screen "0012_Pump Setting" 1280x800, template "Navigation"
   on GenerateScreen: SetBit("DB613_Komponent_State_Read"); SetBit("DB608_PV_Metering_Read")
   Button "Button_1" at 133,154 size 561x639; TextOff 'Text'
   TextField "Text field_1" at 170,166 size 134x25; Text 'Pump enable:'
   TextField "Text field_2" at 170,199 size 128x25; Text 'Machine No.:'
   TextField "Text field_3" at 170,231 size 90x25; Text 'Daytank:'
   TextField "Text field_4" at 170,296 size 65x25; Text 'Name:'
   TextField "Text field_5" at 170,326 size 156x25; Text 'Pulse per. Liter:'
   TextField "Text field_7" at 170,357 size 196x25; Text 'Adjustm. time [ms]:'
   IOField "Pump_Pulse_Perliter" at 453,323 size 166x30; Authorization "User administration"; FormatPattern 99999.999
      ProcessValue <- "DB753_MeteringPump_Pump{0}_Pulse_per_liter"
   TextField "Text field_8" at 170,550 size 82x25; Text 'Control:'
   TextField "Text field_9" at 170,582 size 146x25; Text 'Feeding Pump:'
   TextField "Text field_10" at 170,617 size 114x25; Text 'Edge Filter:'
   TextField "Text field_11" at 170,652 size 181x25; Text 'Cooling / Heating:'
   TextField "Text field_12" at 170,687 size 192x25; Text 'Deselection Enable:'
   TextField "Text field_13" at 170,722 size 302x25; Text 'With min Temperature Release:'
   TextField "Text field_14" at 170,757 size 167x25; Text 'With flow factor:'
   IOField "I/O field_2" at 453,354 size 166x30; Authorization "User administration"; FormatPattern 99999.999
      ProcessValue <- "PN_FlowRate_Component{0}_FlowC_F_GeneralParameters_Data_Nachstellzeit"
   IOField "I/O field_3" at 453,385 size 166x30; Authorization "User administration"; FormatPattern 999.9
      ProcessValue <- "DB753_MeteringPump_Pump{0}_MaxFlowLiter"
   IOField "I/O field_4" at 551,196 size 69x30; Authorization "User administration"; FormatPattern 999
      ProcessValue <- "DB753_MeteringPump_Pump{0}_MachineNumber"
   IOField "I/O field_5" at 551,228 size 69x30; Authorization "User administration"; FormatPattern 9999
      ProcessValue <- "DB753_MeteringPump_Pump{0}_TankNo"
   Button "Check_Pump_Enable" at 575,161 size 45x30; TextOff 'Text'; PictureOff "download"; PictureList "Check_Uncheck"
      ProcessValue <- "DB753_MeteringPump_Pump{0}_Pump_Active"
      on Click: InvertBit("DB753_MeteringPump_Pump{0}_Pump_Active")
   Button "Check_Pump_WithFeedingPump" at 573,579 size 45x30; TextOff 'Text'; PictureOff "download"; PictureList "Check_Uncheck"
      ProcessValue <- "DB753_MeteringPump_Pump{0}_WithFeedPump"
      on Click: InvertBit("DB753_MeteringPump_Pump{0}_WithFeedPump")
   Button "Check_Pump_WithEdgeFilter" at 573,614 size 45x30; TextOff 'Text'; PictureOff "download"; PictureList "Check_Uncheck"
      ProcessValue <- "DB753_MeteringPump_Pump{0}_WithEdgeFilter"
      on Click: InvertBit("DB753_MeteringPump_Pump{0}_WithEdgeFilter")
   Button "Check_Pump_CoolingHeating" at 573,649 size 45x30; TextOff 'Text'; PictureOff "download"; PictureList "Check_Uncheck"
      ProcessValue <- "DB753_MeteringPump_Pump{0}_WithHeating"
      on Click: InvertBit("DB753_MeteringPump_Pump{0}_WithHeating")
   Button "Check_Pump_Deselection_Ena" at 573,684 size 45x30; TextOff 'Text'; PictureOff "download"; PictureList "Check_Uncheck"
      ProcessValue <- "DB753_MeteringPump_Pump{0}_PumDeselectionEnable"
      on Click: InvertBit("DB753_MeteringPump_Pump{0}_PumDeselectionEnable")
   Button "Check_Pump_WithMinTempRelease" at 573,719 size 45x30; TextOff 'Text'; PictureOff "download"; PictureList "Check_Uncheck"
      ProcessValue <- "DB753_MeteringPump_Pump{0}_WithMinTempRelease"
      on Click: InvertBit("DB753_MeteringPump_Pump{0}_WithMinTempRelease")
   Button "Check_Pump_WithFlowFactor" at 573,754 size 45x30; TextOff 'Text'; PictureOff "download"; PictureList "Check_Uncheck"
      ProcessValue <- "DB753_MeteringPump_Pump{0}_WithFlowFactor"
      on Click: InvertBit("DB753_MeteringPump_Pump{0}_WithFlowFactor")
   Button "b_Incress_Pump_Setting" at 785,104 size 46x32; TextOff 'Text'; PictureOff "right arrow"
      on Click: function_dd21b452("DB613_Komponent_State_ReadDeviceNo", 1); function_dd21b452("DB612_Tank_State.ReadDeviceNo", 1)
   Button "b_Decress_Pump_Setting" at 273,104 size 46x32; TextOff 'Text'; PictureOff "left arrow"
      on Click: function_b9b71300("DB613_Komponent_State_ReadDeviceNo", 1); function_b9b71300("DB612_Tank_State.ReadDeviceNo", 1)
   Button "b_Pump_Control" at 503,547 size 45x30; TextOff 'Text'; PictureOff "obeng"
      on Click: SetTag("Control", 1)
   Button "b_Pump_Feeding_Pump" at 503,579 size 45x30; TextOff 'Text'; PictureOff "obeng"
      on Click: SetTag("Control", 2)
      Visibility <- "DB753_MeteringPump_Pump{0}_WithFeedPump"
   Button "b_Pump_EdgeFilter" at 503,615 size 45x30; TextOff 'Text'; PictureOff "obeng"
      on Click: SetTag("Control", 3)
      Visibility <- "DB753_MeteringPump_Pump{0}_WithEdgeFilter"
   Button "b_Pump_CoolingHeating" at 503,651 size 45x30; TextOff 'Text'; PictureOff "obeng"
      on Click: SetTag("Control", 4)
      Visibility <- "DB753_MeteringPump_Pump{0}_WithHeating"
   IOField "I/O field_6" at 453,293 size 166x30; Authorization "User administration"; FormatPattern ??????????
      ProcessValue <- "DB753_MeteringPump_Pump{0}_Name"
   IOField "I/O field_7" at 382,261 size 236x30; Authorization "User administration"; FormatPattern ??????????
      ProcessValue <- "DB753_MeteringPump_Pump{0}_Name"
   IOField "I/O field_8" at 453,417 size 166x30; Authorization "User administration"; FormatPattern 999.9
      ProcessValue <- "DB753_MeteringPump_Pump{0}_MinFlowPercent"
   IOField "I/O field_9" at 453,449 size 166x30; Authorization "User administration"; FormatPattern 999.9
      ProcessValue <- "DB753_MeteringPump_Pump{0}_MaxFlowPercent"
   IOField "I/O field_10" at 453,479 size 166x30; Authorization "User administration"; FormatPattern 99999.99
      ProcessValue <- "DB613_Komponent_State_FlowPumpMin{0}"
   IOField "I/O field_11" at 453,511 size 166x30; Authorization "User administration"; FormatPattern 99999.99
      ProcessValue <- "DB613_Komponent_State_FlowPumpMax{0}"
   TextField "Text field_20" at 170,388 size 227x25; Text 'Pump quantity [l/min]:'
   TextField "Text field_21" at 170,420 size 142x25; Text 'Min. Flow[%]:'
   TextField "Text field_22" at 170,452 size 146x25; Text 'Max. Flow[%]:'
   TextField "Text field_23" at 170,482 size 154x25; Text 'Min. Flow[g/s]:'
   TextField "Text field_24" at 170,514 size 158x25; Text 'Max. Flow[g/s]:'
   IOField "I/O field_43" at 326,104 size 451x32; FormatPattern ????????????????????
      ProcessValue <- "DB753_MeteringPump_Pump{0}_Name"
      Appearance <- "DB702_Tank_Value_Tank{0}_Color"
   Button "Button_19" at 856,366 size 159x83; TextOff 'Text'; PictureOff "motor_2"; PictureList "pump"
      ProcessValue <- "DB613_Komponent_State_ReadDeviceNo"
      Visibility <- "DB753_MeteringPump_Pump{0}_Pump_Active"
   GraphicView "Graphic view_1" at 763,170 size 81x40; Picture "motor2"
      Visibility <- "DB753_MeteringPump_Pump{0}_WithFeedPump"
   GraphicView "Graphic view_2" at 715,254 size 125x120; Picture "heatHP"
      Visibility <- "DB753_MeteringPump_Pump{0}_WithHeating"
   GraphicView "Graphic view_5" at 1047,261 size 58x89; Picture "heatLP"
      Visibility <- "DB753_MeteringPump_Pump{0}_WithLPHeatExchanger"
   GraphicView "Graphic view_7" at 977,170 size 67x93; Picture "edgefilter"
      Visibility <- "DB753_MeteringPump_Pump{0}_WithEdgeFilter"
   GraphicView "Graphic view_9" at 1112,275 size 39x75; Picture "Graphic_14"
      Visibility <- "DB753_MeteringPump_Pump{0}_WithFischerValveLP"
   GraphicView "Graphic view_10" at 801,275 size 39x75; Picture "Graphic_14"
      Visibility <- "DB753_MeteringPump_Pump{0}_WithFischerValveHP"
   Button "Button_8" at 720,466 size 437x286; TextOff 'Text'
      Visibility <- "Control"
   TextField "Text field_15" at 742,497 size 169x30; Text 'Control Pump:'
      Visibility <- "Control"
   TextField "Text field_16" at 742,573 size 91x25; Text 'With FC :'
      Visibility <- "Control"
   TextField "Text field_17" at 742,617 size 104x25; Text 'Controlled'
      Visibility <- "Control"
   TextField "Text field_18" at 742,661 size 73x25; Text '2 Point'
      Visibility <- "Control"
   TextField "Text field_19" at 940,617 size 101x25; Text 'Regulated'
      Visibility <- "Control"
   Button "Check_Pump_ControlPump_WithFc" at 862,570 size 45x30; TextOff 'Text'; PictureOff "download"; PictureList "Check_Uncheck"
      ProcessValue <- "DB753_MeteringPump_Pump{0}_WithFC"
      Visibility <- "Control"
      on Click: InvertBit("DB753_MeteringPump_Pump{0}_WithFC")
   Button "Check_Pump_ControlPump_Controlled" at 862,614 size 45x30; TextOff 'Text'; PictureOff "download"; PictureList "Check_Uncheck"
      Visibility <- "Control"
      ProcessValue <- "DB753_MeteringPump_Pump{0}_WithFlowControl"
      on Click: InvertBit("DB753_MeteringPump_Pump{0}_WithFlowControl")
   Button "Check_Pump_ControlPump_2Point" at 862,658 size 45x30; TextOff 'Text'; PictureOff "download"; PictureList "Check_Uncheck"
      ProcessValue <- "DB753_MeteringPump_Pump{0}_With_2Point"
      Visibility <- "Control"
      on Click: InvertBit("DB753_MeteringPump_Pump{0}_With_2Point")
   Button "Check_Pump_ControlPump_Regulated" at 1057,614 size 45x30; TextOff 'Text'; PictureOff "download"; PictureList "Check_Uncheck"
      Visibility <- "Control"
      ProcessValue <- "DB753_MeteringPump_Pump{0}_WithoutFlowControl"
      on Click: InvertBit("DB753_MeteringPump_Pump{0}_WithoutFlowControl")
   Button "b_Pump_Close_ControlPump" at 1101,470 size 51x41; TextOff 'Text'; PictureOff "images (1)"
      Visibility <- "Control"
      on Click: SetTag("Control", 0)
   Button "Button_2" at 720,466 size 437x286; TextOff 'Text'
      Visibility <- "Control"
   TextField "Text field_6" at 758,496 size 173x30; Text 'Feeding Pump:'
      Visibility <- "Control"
   TextField "Text field_25" at 794,559 size 78x25; Text 'With FC'
      Visibility <- "Control"
   TextField "Text field_26" at 794,609 size 157x25; Text 'No pressure ctr.'
      Visibility <- "Control"
   TextField "Text field_27" at 794,657 size 72x25; Text 'Bypass'
      Visibility <- "Control"
   TextField "Text field_28" at 1023,559 size 125x25; Text 'Pressure ctr.'
      Visibility <- "Control"
   Button "Check_Pump_FP_WithFC" at 738,556 size 45x30; TextOff 'Text'; PictureOff "download"; PictureList "Check_Uncheck"
      Visibility <- "Control"
      on Click: InvertBit("DB751_auxiliaryDriveMetering_FeedingPump{0}_Config_WithFC")
      ProcessValue <- "DB751_auxiliaryDriveMetering_FeedingPump{0}_Config_WithFC"
   Button "Check_Pump_FP_NoPressCtr" at 738,606 size 45x30; TextOff 'Text'; PictureOff "download"; PictureList "Check_Uncheck"
      Visibility <- "Control"
      on Click: InvertBit("DB751_auxiliaryDriveMetering_FeedingPump{0}_Config_Without_PresControl")
      ProcessValue <- "DB751_auxiliaryDriveMetering_FeedingPump{0}_Config_Without_PresControl"
   Button "Check_Pump_FP_Bypass" at 738,654 size 45x30; TextOff 'Text'; PictureOff "download"; PictureList "Check_Uncheck"
      Visibility <- "Control"
      on Click: InvertBit("DB751_auxiliaryDriveMetering_FeedingPump{0}_Config_Bypass")
      ProcessValue <- "DB751_auxiliaryDriveMetering_FeedingPump{0}_Config_Bypass"
   Button "Check_Pump_FP_PressureCtr" at 963,556 size 45x30; TextOff 'Text'; PictureOff "download"; PictureList "Check_Uncheck"
      Visibility <- "Control"
      on Click: InvertBit("DB751_auxiliaryDriveMetering_FeedingPump{0}_Config_With_PresControl")
      ProcessValue <- "DB751_auxiliaryDriveMetering_FeedingPump{0}_Config_With_PresControl"
   Button "b_Close_Pump_FeddingPump" at 1101,469 size 51x41; TextOff 'Text'; PictureOff "images (1)"
      Visibility <- "Control"
      on Click: SetTag("Control", 0)
   TextField "Text field_29" at 794,705 size 154x25; Text 'Manual Switch?'
      Visibility <- "Control"
   Button "Check_Pump_FP_ManualSwtch?" at 738,702 size 45x30; TextOff 'Text'; PictureOff "download"; PictureList "Check_Uncheck"
      Visibility <- "Control"
      on Click: InvertBit("DB751_auxiliaryDriveMetering_FeedingPump{0}_Config_ManualSwitchON")
      ProcessValue <- "DB751_auxiliaryDriveMetering_FeedingPump{0}_Config_ManualSwitchON"
   TextField "Text field_30" at 1023,609 size 64x25; Text 'Filling'
      Visibility <- "Control"
   Button "Check-Pump_FP_Filling" at 963,606 size 45x30; TextOff 'Text'; PictureOff "download"; PictureList "Check_Uncheck"
      Visibility <- "Control"
      on Click: InvertBit("DB751_auxiliaryDriveMetering_FeedingPump{0}_Config_Filling")
      ProcessValue <- "DB751_auxiliaryDriveMetering_FeedingPump{0}_Config_Filling"
   Button "Button_11" at 720,466 size 437x286; TextOff 'Text'
      Visibility <- "Control"
   TextField "Text field_31" at 754,496 size 136x30; Text 'Edge Filter:'
      Visibility <- "Control"
   TextField "Text field_32" at 810,559 size 111x25; Text 'With Motor'
      Visibility <- "Control"
   TextField "Text field_33" at 810,609 size 72x25; Text 'Double'
      Visibility <- "Control"
   TextField "Text field_35" at 1023,609 size 125x25; Text 'Pressure ctr.'
      Visibility <- "Control"
   Button "Check_Pump_EF_WithMotor" at 754,556 size 45x30; TextOff 'Text'; PictureOff "download"; PictureList "Check_Uncheck"
      Visibility <- "Control"
      on Click: InvertBit("DB751_auxiliaryDriveMetering_EdgeFilter{0}_Config_Driven")
      ProcessValue <- "DB751_auxiliaryDriveMetering_EdgeFilter{0}_Config_Driven"
   Button "Check_Pump_EF_Double" at 754,606 size 45x30; TextOff 'Text'; PictureOff "download"; PictureList "Check_Uncheck"
      Visibility <- "Control"
      on Click: InvertBit("DB751_auxiliaryDriveMetering_EdgeFilter{0}_Config_Double")
      ProcessValue <- "DB751_auxiliaryDriveMetering_EdgeFilter{0}_Config_Double"
   Button "Check_Pump_EF_Pressurectr" at 963,606 size 45x30; TextOff 'Text'; PictureOff "download"; PictureList "Check_Uncheck"
      Visibility <- "Control"
      on Click: InvertBit("DB751_auxiliaryDriveMetering_FeedingPump{0}_Config_With_PresControl")
      ProcessValue <- "DB751_auxiliaryDriveMetering_FeedingPump{0}_Config_With_PresControl"
   Button "b_Close_Pump_EdgeFilter_Close" at 1101,469 size 51x41; TextOff 'Text'; PictureOff "images (1)"
      Visibility <- "Control"
      on Click: SetTag("Control", 0)
   Button "Button_13" at 720,465 size 437x286; TextOff 'Text'
      Visibility <- "Control"
   TextField "Text field_34" at 758,496 size 222x30; Text 'Cooling / Heating :'
      Visibility <- "Control"
   TextField "Text field_36" at 794,559 size 83x25; Text 'Exhause'
      Visibility <- "Control"
   TextField "Text field_37" at 794,609 size 132x25; Text 'LP Exchanger'
      Visibility <- "Control"
   TextField "Text field_38" at 794,657 size 135x25; Text 'HP Exchanger'
      Visibility <- "Control"
   TextField "Text field_39" at 1023,559 size 129x25; Text 'Fischer valve'
      Visibility <- "Control"
   Button "Check_Pump_CH_Exhause" at 738,556 size 45x30; TextOff 'Text'; PictureOff "download"; PictureList "Check_Uncheck"
      Visibility <- "Control"
      ProcessValue <- "DB753_MeteringPump_Pump{0}_WithExhauseSystem"
      on Click: InvertBit("DB753_MeteringPump_Pump{0}_WithExhauseSystem")
   Button "Check_Pump_CH_LPExchanger" at 738,606 size 45x30; TextOff 'Text'; PictureOff "download"; PictureList "Check_Uncheck"
      Visibility <- "Control"
      ProcessValue <- "DB753_MeteringPump_Pump{0}_WithLPHeatExchanger"
      on Click: InvertBit("DB753_MeteringPump_Pump{0}_WithLPHeatExchanger")
   Button "Check_Pump_CH_HPExchanger" at 738,654 size 45x30; TextOff 'Text'; PictureOff "download"; PictureList "Check_Uncheck"
      Visibility <- "Control"
      on Click: InvertBit("DB753_MeteringPump_Pump{0}_WithHeating")
      ProcessValue <- "DB753_MeteringPump_Pump{0}_WithHeating"
   Button "Check_Pump_CH_FischerLP" at 963,556 size 45x30; TextOff 'Text'; PictureOff "download"; PictureList "Check_Uncheck"
      Visibility <- "Control"
      on Click: InvertBit("DB753_MeteringPump_Pump{0}_WithFischerValveLP")
      ProcessValue <- "DB753_MeteringPump_Pump{0}_WithFischerValveLP"
   TextField "Text field_40" at 794,705 size 46x25; Text 'Pipe'
      Visibility <- "Control"
   Button "Check_Pump_CH_Pipe" at 738,702 size 45x30; TextOff 'Text'; PictureOff "download"; PictureList "Check_Uncheck"
      Visibility <- "Control"
      on Click: InvertBit("DB753_MeteringPump_Pump{0}_With_2Point")
      ProcessValue <- "DB753_MeteringPump_Pump{0}_With_2Point"
   TextField "Text field_41" at 1023,609 size 129x25; Text 'Fischer valve'
      Visibility <- "Control"
   Button "Check_Pump_CH_FischerHP" at 963,606 size 45x30; TextOff 'Text'; PictureOff "download"; PictureList "Check_Uncheck"
      Visibility <- "Control"
      on Click: InvertBit("DB753_MeteringPump_Pump{0}_WithFischerValveHP")
      ProcessValue <- "DB753_MeteringPump_Pump{0}_WithFischerValveHP"
   Button "b_Close_Pump_CH" at 1101,469 size 51x41; TextOff 'Text'; PictureOff "images (1)"
      on Press: SetTag("Control", 0)
      Visibility <- "Control"

screen "0007_Tank Setting" 1280x800, template "Navigation"
   on GenerateScreen: SetBit("DB612_Tank_State.Read")
   Button "Tank_Bg" at 118,165 size 535x569; TextOff 'Text'
      Visibility <- "DB702_Tank_Value_Tank{0}_Deselected"
   TextField "Text field_1" at 166,212 size 65x25; Text 'Name:'
      Visibility <- "DB702_Tank_Value_Tank{0}_Deselected"
   TextField "Text field_2" at 166,245 size 82x25; Text 'Display:'
      Visibility <- "DB702_Tank_Value_Tank{0}_Deselected"
   TextField "Text field_3" at 166,310 size 84x25; Text 'Density:'
      Visibility <- "DB702_Tank_Value_Tank{0}_Deselected"
   TextField "Text field_4" at 166,348 size 122x25; Text 'Filling level:'
      Visibility <- "DB702_Tank_Value_Tank{0}_Deselected"
   TextField "Text field_5" at 166,382 size 71x25; Text 'Filling:'
      Visibility <- "DB702_Tank_Value_Tank{0}_Deselected"
   TextField "Text field_6" at 166,416 size 114x25; Text 'Nucleation:'
      Visibility <- "DB702_Tank_Value_Tank{0}_Deselected"
   TextField "Text field_7" at 166,450 size 186x25; Text 'Tempering control:'
      Visibility <- "DB702_Tank_Value_Tank{0}_Deselected"
   TextField "Text field_8" at 166,484 size 86x25; Text 'Vacuum:'
      Visibility <- "DB702_Tank_Value_Tank{0}_Deselected"
   TextField "Text field_9" at 166,518 size 101x25; Text 'Emptying:'
      Visibility <- "DB702_Tank_Value_Tank{0}_Deselected"
   TextField "Text field_10" at 166,552 size 142x25; Text 'Barrel station:'
      Visibility <- "DB702_Tank_Value_Tank{0}_Deselected"
   TextField "Text field_11" at 166,586 size 122x25; Text 'Tank stirrer:'
      Visibility <- "DB702_Tank_Value_Tank{0}_Deselected"
   TextField "Text field_12" at 166,620 size 140x25; Text 'Force stirring:'
      Visibility <- "DB702_Tank_Value_Tank{0}_Deselected"
   TextField "Text field_13" at 166,654 size 141x25; Text 'Deselect tank:'
      Visibility <- "DB702_Tank_Value_Tank{0}_Deselected"
   TextField "Text field_14" at 166,688 size 196x25; Text 'Pentane equipment:'
      Visibility <- "DB702_Tank_Value_Tank{0}_Deselected"
   IOField "Tank_Density" at 425,307 size 100x30; Authorization "User administration"; FormatPattern 99999
      ProcessValue <- "DB702_Tank_Value.Tank[0].Density"
      Visibility <- "DB702_Tank_Value_Tank{0}_Deselected"
   TextField "Text field_16" at 546,311 size 46x25; Text 'g/l'
      Visibility <- "DB702_Tank_Value_Tank{0}_Deselected"
   Button "b_FillingLevel" at 539,343 size 45x30; TextOff 'Text'; PictureOff "obeng"
      Visibility <- "DB702_Tank_Value_Tank{0}_Deselected"
      on Click: SetTag("Control2", 1)
   Button "b_Filling" at 539,378 size 45x30; TextOff 'Text'; PictureOff "obeng"
      Visibility <- "DB702_Tank_Value_Tank{0}_Deselected"
      on Click: SetTag("Control2", 2)
   Button "b_TemperingControl" at 539,447 size 45x30; TextOff 'Text'; PictureOff "obeng"
      Visibility <- "DB702_Tank_Value_Tank{0}_Deselected"
      on Click: SetTag("Control2", 3)
   Button "b_BarrelStation" at 539,548 size 45x30; TextOff 'Text'; PictureOff "obeng"
      Visibility <- "DB702_Tank_Value_Tank{0}_Deselected"
      on Click: SetTag("Control2", 4)
   Button "b_TankStirree" at 539,581 size 45x30; TextOff 'Text'; PictureOff "obeng"
      Visibility <- "DB702_Tank_Value_Tank{0}_Deselected"
      on Click: SetTag("Control2", 5)
   Button "b_ForceStrirring" at 539,617 size 45x30; TextOff 'Text'; PictureOff "obeng"
      Visibility <- "DB702_Tank_Value_Tank{0}_Deselected"
      on Click: SetTag("Control2", 6)
   IOField "I/O field_6" at 425,210 size 166x30; Authorization "User administration"; FormatPattern ??????????
      ProcessValue <- "DB702_Tank_Value_Tank{0}_Name"
      Visibility <- "DB702_Tank_Value_Tank{0}_Deselected"
   Button "Check_Nucleation" at 538,414 size 45x30; TextOff 'Text'; PictureOff "download"; PictureList "Check_Uncheck"
      ProcessValue <- "DB702_Tank_Value_Tank{0}_With_Nucleation"
      Visibility <- "DB702_Tank_Value_Tank{0}_Deselected"
      on Click: InvertBit("DB702_Tank_Value_Tank{0}_With_Nucleation")
   Button "Check_WithVacum" at 538,482 size 45x30; TextOff 'Text'; PictureOff "download"; PictureList "Check_Uncheck"
      ProcessValue <- "DB702_Tank_Value_Tank{0}_With_Vacuum"
      Visibility <- "DB702_Tank_Value_Tank{0}_Deselected"
      on Click: InvertBit("DB702_Tank_Value_Tank{0}_With_Vacuum")
   Button "Check_Emptyting" at 538,516 size 45x30; TextOff 'Text'; PictureOff "download"; PictureList "Check_Uncheck"
      Visibility <- "DB702_Tank_Value_Tank{0}_Deselected"
      on Click: InvertBit("DB702_Tank_Value_Tank{0}_With_Drain")
      ProcessValue <- "DB702_Tank_Value_Tank{0}_With_Drain"
   Button "Check_Deselect_Tank" at 538,649 size 45x30; TextOff 'Text'; PictureList "Check_Uncheck"; PictureOff "images (7)"
      on Click: InvertBit("DB702_Tank_Value_Tank{0}_Existing")
      ProcessValue <- "DB702_Tank_Value_Tank{0}_Existing"
   Button "Check_Pentane" at 538,683 size 45x30; TextOff 'Text'; PictureOff "download"; PictureList "Check_Uncheck"
      ProcessValue <- "DB702_Tank_Value_Tank{0}_With_Filling_Pentane"
      Visibility <- "DB702_Tank_Value_Tank{0}_Deselected"
      on Click: InvertBit("DB702_Tank_Value_Tank{0}_With_Filling_Pentane")
   Button "b_Increess_Tank_Setting" at 788,104 size 46x32; TextOff 'Text'; PictureOff "right arrow"
      on Click: function_dd21b452("DB612_Tank_State.ReadDeviceNo", 1)
   Button "b_Decress_Tank_Setting" at 269,104 size 46x32; TextOff 'Text'; PictureOff "left arrow"
      on Click: function_b9b71300("DB612_Tank_State.ReadDeviceNo", 1)
   IOField "I/O field_43" at 326,104 size 451x32; FormatPattern ????????????????????
      ProcessValue <- "DB702_Tank_Value_Tank{0}_Name"
      Appearance <- "DB702_Tank_Value_Tank{0}_Color"
   GraphicIOField "Graphic I/O field_1" at 425,249 size 166x50; PictureList "Color"; Authorization "User administration"
      ProcessValue <- "DB702_Tank_Value_Tank{0}_Color"
      Visibility <- "DB702_Tank_Value_Tank{0}_Deselected"
   GraphicView "Graphic view_2" at 760,560 size 129x217; Picture "tank"
   Bar "Bar_1" at 809,585 size 33x143; MinimumValue 0; MaximumValue 100
      ProcessValue <- "DB602_PV_Tank_Tank{0}_Level_PV_ActV_Value"
      Visibility <- "DB702_Tank_Value_Tank{0}_With_Level_Probe"
   GraphicIOField "Graphic I/O field_2" at 772,592 size 25x20; PictureList "Tank_Sensor"
      Visibility <- "DB702_Tank_Value_Tank{0}_With_Level_3Liq"
      ProcessValue <- "DB612_Tank_State_Tank{0}_Stop_Level_Filling"
   GraphicIOField "Graphic I/O field_3" at 772,630 size 25x20; PictureList "Tank_Sensor"
      Visibility <- "DB702_Tank_Value_Tank{0}_With_Level_4Liq"
      ProcessValue <- "DB612_Tank_State_Tank{0}_Start_Level_Filling"
   GraphicIOField "Smin" at 772,709 size 25x20; PictureList "Tank_Sensor"
      Visibility <- "DB702_Tank_Value_Tank{0}_With_Level_SMin"
      ProcessValue <- "DB612_Tank_State_Tank{0}_Min_Level"
   GraphicIOField "Smax" at 848,592 size 25x20; PictureList "Tank_Sensor"
      Visibility <- "DB702_Tank_Value_Tank{0}_With_Level_SMax"
      ProcessValue <- "DB612_Tank_State_Tank{0}_Max_Level"
   GraphicIOField "Graphic I/O field_6" at 890,560 size 25x20; PictureList "Tank_Sensor"
      Visibility <- "DB702_Tank_Value_Tank{0}_With_Filling_Switch"
      ProcessValue <- "DB612_Tank_State_Tank{0}_Max_Level"
   GraphicView "Graphic view_3" at 888,592 size 32x45; Picture "Graphic_7"
      Visibility <- "DB702_Tank_Value_Tank{0}_With_Filling_Valve"
   GraphicView "Graphic view_4" at 936,592 size 32x45; Picture "Graphic_7"
      Visibility <- "DB702_Tank_Value_Tank{0}_With_Filling_2Valve"
   GraphicIOField "Graphic I/O field_7" at 936,560 size 25x20; PictureList "Tank_Sensor"
      Visibility <- "DB702_Tank_Value_Tank{0}_With_Filling_Switch"
      ProcessValue <- "DB612_Tank_State_Tank{0}_Max_Level"
   GraphicView "Graphic view_5" at 888,696 size 32x45; Picture "Graphic_7"
      Visibility <- "DB702_Tank_Value_Tank{0}_With_Filling_ShutDown"
   Rectangle "Rectangle_1" at 883,552 size 40x40
      Visibility <- "DB702_Tank_Value_Tank{0}_With_Filling_Valve"
   Rectangle "Rectangle_2" at 928,550 size 45x40
      Visibility <- "DB702_Tank_Value_Tank{0}_With_Filling_2Valve"
   GraphicView "Graphic view_7" at 1000,736 size 32x45; Picture "Graphic_14"
      Visibility <- "DB702_Tank_Value_Tank{0}_With_Tempering_WTmitFischer"
   GraphicView "Graphic view_8" at 696,656 size 72x117; Picture "HeaterBackFL"
      Visibility <- "DB702_Tank_Value_Tank{0}_With_Tempering_WTRL"
   GraphicView "Graphic view_9" at 804,755 size 41x35; Picture "HEATER"
      Visibility <- "DB702_Tank_Value_Tank{0}_With_Tempering_Heizung"
   GraphicView "Graphic view_10" at 936,712 size 60x77; Picture "heatLP"
      Visibility <- "DB702_Tank_Value_Tank{0}_With_Tempering_WTVL"
   GraphicView "Graphic view_11" at 1040,616 size 75x86; Picture "Graphic_16"
      Visibility <- "DB702_Tank_Value_Tank{0}_With_BarelStation"
   GraphicView "Graphic view_1" at 800,524 size 53x54; Picture "Graphic_17"
      Visibility <- "DB702_Tank_Value_Tank{0}_With_Agitator"
   GraphicView "Graphic view_12" at 726,528 size 26x38; Picture "Graphic_18"
      Visibility <- "DB702_Tank_Value_Tank{0}_With_Agitator_Converter"
   GraphicIOField "Graphic I/O field_15" at 732,584 size 34x30; PictureList "Valve_Tank"
      Visibility <- "DB702_Tank_Value_Tank{0}_With_Tempering_VKaltwasser"
      ProcessValue <- "Internal_Tank_"
   GraphicIOField "Graphic I/O field_8" at 693,748 size 34x30; PictureList "Valve_Tank"
      ProcessValue <- "Internal_Tank_"
      Visibility <- "DB702_Tank_Value_Tank{0}_With_Tempering_WTRL"
   GraphicView "Graphic view_13" at 886,527 size 35x29; Picture "startfilling"
      Visibility <- "DB612_Tank_State_Tank{0}_Filling_Start"
   GraphicIOField "3Level Smax" at 848,592 size 25x20; PictureList "Tank_Sensor"
      ProcessValue <- "DB612_Tank_State_Tank{0}_Max_Level"
      Visibility <- "DB702_Tank_Value_Tank{0}_With_Level_3Liq"
   GraphicIOField "3Level Smin" at 772,709 size 25x20; PictureList "Tank_Sensor"
      ProcessValue <- "DB612_Tank_State_Tank{0}_Min_Level"
      Visibility <- "DB702_Tank_Value_Tank{0}_With_Level_3Liq"
   GraphicIOField "4Level Liq" at 772,592 size 25x20; PictureList "Tank_Sensor"
      ProcessValue <- "DB612_Tank_State_Tank{0}_Stop_Level_Filling"
      Visibility <- "DB702_Tank_Value_Tank{0}_With_Level_4Liq"
   GraphicIOField "4Level Smin" at 772,709 size 25x20; PictureList "Tank_Sensor"
      ProcessValue <- "DB612_Tank_State_Tank{0}_Min_Level"
      Visibility <- "DB702_Tank_Value_Tank{0}_With_Level_4Liq"
   GraphicIOField "4Level Smax" at 848,592 size 25x20; PictureList "Tank_Sensor"
      ProcessValue <- "DB612_Tank_State_Tank{0}_Max_Level"
      Visibility <- "DB702_Tank_Value_Tank{0}_With_Level_4Liq"
   GraphicView "Graphic view_6" at 888,592 size 32x45; Picture "Graphic_7"
      Visibility <- "DB702_Tank_Value_Tank{0}_With_Filling_ShutDown"
   GraphicView "Alarm Indicator Tank2_1" at 761,534 size 28x25; Picture "AlarmState2"
      Visibility <- "DB612_Tank_State_Agitator{0}_FLT_Exist"
   Button "b_Tank2_1" at 753,530 size 48x32; TextOff 'Text'
      on Press: ActivateScreen("0024_ActualFaults", 0); SetTag("Alarm_Filter_Tag", 4)
      ObjectEnable <- "DB612_Tank_State_FaultExists{2}"
   GraphicView "Graphic view_14" at 766,498 size 35x29; Picture "startfilling"
      Visibility <- "DB612_Tank_State_Agitator{0}_Run"
   GraphicIOField "Graphic I/O field_13" at 932,532 size 25x20; PictureList "Tank_Sensor"
      ProcessValue <- "DB612_Tank_State_Tank{0}_Max_Level"
      Visibility <- "DB702_Tank_Value_Tank{0}_With_Filling_Switch"
   Button "FLD POPUP" at 692,165 size 451x280; TextOff 'Text'
      Visibility <- "Control2"
   TextField "Text field_17" at 766,249 size 81x25; Text 'Existing'
      Visibility <- "Control2"
   TextField "Text field_18" at 766,296 size 143x25; Text '3 Level Switch'
      Visibility <- "Control2"
   TextField "Text field_19" at 766,343 size 116x25; Text 'Level Probe'
      Visibility <- "Control2"
   TextField "Text field_20" at 1002,249 size 127x25; Text '+ Super Min.'
      Visibility <- "Control2"
   TextField "Text field_21" at 1002,296 size 143x25; Text '4 Level Switch'
      Visibility <- "Control2"
   TextField "Text field_22" at 1002,343 size 131x25; Text '+ Super Max.'
      Visibility <- "Control2"
   TextField "Text field_15" at 719,194 size 240x30; Text 'Filling Level Display:'
      Visibility <- "Control2"
   Button "Check_Tank_FLD_Existing" at 711,246 size 45x30; TextOff 'Text'; PictureOff "download"; PictureList "Check_Uncheck"
      Visibility <- "Control2"
      on Click: InvertBit("DB702_Tank_Value_Tank{0}_With_Level")
      ProcessValue <- "DB702_Tank_Value_Tank{0}_With_Level"
   Button "Check_Tank_FLD_3LevelSwitch" at 711,293 size 45x30; TextOff 'Text'; PictureOff "download"; PictureList "Check_Uncheck"
      Visibility <- "Control2"
      ProcessValue <- "DB702_Tank_Value_Tank{0}_With_Level_3Liq"
      on Click: InvertBit("DB702_Tank_Value_Tank{0}_With_Level_3Liq")
   Button "Check_Tank_FLD_LevelProbe" at 711,340 size 45x30; TextOff 'Text'; PictureOff "download"; PictureList "Check_Uncheck"
      Visibility <- "Control2"
      ProcessValue <- "DB702_Tank_Value_Tank{0}_With_Level_Probe"
      on Click: InvertBit("DB702_Tank_Value_Tank{0}_With_Level_Probe")
   Button "Check_Tank_FLD_Smin" at 948,246 size 45x30; TextOff 'Text'; PictureOff "download"; PictureList "Check_Uncheck"
      Visibility <- "Control2"
      ProcessValue <- "DB702_Tank_Value_Tank{0}_With_Level_SMin"
      on Click: InvertBit("DB702_Tank_Value_Tank{0}_With_Level_SMin")
   Button "Check_Tank_FLD_4LevelSwitch" at 948,293 size 45x30; TextOff 'Text'; PictureOff "download"; PictureList "Check_Uncheck"
      Visibility <- "Control2"
      ProcessValue <- "DB702_Tank_Value_Tank{0}_With_Level_4Liq"
      on Click: InvertBit("DB702_Tank_Value_Tank{0}_With_Level_4Liq")
   Button "Check_Tank_FLD_Smax" at 948,340 size 45x30; TextOff 'Text'; PictureOff "download"; PictureList "Check_Uncheck"
      Visibility <- "Control2"
      ProcessValue <- "DB702_Tank_Value_Tank{0}_With_Level_SMax"
      on Click: InvertBit("DB702_Tank_Value_Tank{0}_With_Level_SMax")
   Button "b_Tank_Close_FillingLevelDisplay" at 1087,169 size 51x41; TextOff 'Text'; PictureOff "images (1)"
      Visibility <- "Control2"
      on Click: SetTag("Control2", 0)
   Button "KOF_POPUP" at 692,166 size 451x280; TextOff 'Text'
      Visibility <- "Control2"
   TextField "Text field_23" at 766,250 size 81x25; Text 'Existing'
      Visibility <- "Control2"
   TextField "Text field_24" at 766,297 size 56x25; Text 'Valve'
      Visibility <- "Control2"
   TextField "Text field_25" at 766,344 size 107x25; Text 'Shut down'
      Visibility <- "Control2"
   TextField "Text field_26" at 1002,250 size 140x25; Text 'Containerstat.'
      Visibility <- "Control2"
   TextField "Text field_27" at 1002,297 size 74x25; Text '2 Valve'
      Visibility <- "Control2"
   TextField "Text field_28" at 1002,344 size 120x25; Text 'With Sensor'
      Visibility <- "Control2"
   TextField "Text field_29" at 711,195 size 178x30; Text 'Kind of Filling :'
      Visibility <- "Control2"
   Button "Check_Tank_KOF_Existing" at 711,247 size 45x30; TextOff 'Text'; PictureOff "download"; PictureList "Check_Uncheck"
      Visibility <- "Control2"
      ProcessValue <- "DB702_Tank_Value_Tank{0}_With_Filling"
      on Click: InvertBit("DB702_Tank_Value_Tank{0}_With_Filling")
   Button "Check_Tank_KOF_Valve" at 711,294 size 45x30; TextOff 'Text'; PictureOff "download"; PictureList "Check_Uncheck"
      Visibility <- "Control2"
      ProcessValue <- "DB702_Tank_Value_Tank{0}_With_Filling_Valve"
      on Click: InvertBit("DB702_Tank_Value_Tank{0}_With_Filling_Valve")
   Button "Check_Tank_KOF_Shutdown" at 711,341 size 45x30; TextOff 'Text'; PictureOff "download"; PictureList "Check_Uncheck"
      Visibility <- "Control2"
      ProcessValue <- "DB702_Tank_Value_Tank{0}_With_Filling_ShutDown"
      on Click: InvertBit("DB702_Tank_Value_Tank{0}_With_Filling_ShutDown")
   Button "Check_Tank_KOF_Containerstat" at 948,247 size 45x30; TextOff 'Text'; PictureOff "download"; PictureList "Check_Uncheck"
      Visibility <- "Control2"
      ProcessValue <- "DB702_Tank_Value_Tank{0}_With_ContainerStation"
      on Click: InvertBit("DB702_Tank_Value_Tank{0}_With_ContainerStation")
   Button "Check_Tank_KOF_2Valve" at 948,294 size 45x30; TextOff 'Text'; PictureOff "download"; PictureList "Check_Uncheck"
      Visibility <- "Control2"
      ProcessValue <- "DB702_Tank_Value_Tank{0}_With_Filling_2Valve"
      on Click: InvertBit("DB702_Tank_Value_Tank{0}_With_Filling_2Valve")
   Button "Check_Tank_KOF_WithSensor" at 948,341 size 45x30; TextOff 'Text'; PictureOff "download"; PictureList "Check_Uncheck"
      Visibility <- "Control2"
      ProcessValue <- "DB702_Tank_Value_Tank{0}_With_Filling_Switch"
      on Click: InvertBit("DB702_Tank_Value_Tank{0}_With_Filling_Switch")
   Button "b_Tank_Close_KindFilling" at 1087,170 size 51x41; TextOff 'Text'; PictureOff "images (1)"
      on Press: SetTag("Control2", 0)
      Visibility <- "Control2"
   TextField "Text field_30" at 766,389 size 140x25; Text 'With fill.pump'
      Visibility <- "Control2"
   Button "Check_Tank_KOF_WithFillPump" at 711,386 size 45x30; TextOff 'Text'; PictureOff "download"; PictureList "Check_Uncheck"
      Visibility <- "Control2"
      ProcessValue <- "DB702_Tank_Value_Tank{0}_With_Filling_Pump"
      on Click: InvertBit("DB702_Tank_Value_Tank{0}_With_Filling_Pump")
   TextField "Text field_31" at 1002,390 size 125x25; Text 'With DryRun'
      Visibility <- "Control2"
   Button "Check_Tank_KOF_WithDryRun" at 948,387 size 45x30; TextOff 'Text'; PictureOff "download"; PictureList "Check_Uncheck"
      Visibility <- "Control2"
      ProcessValue <- "DB702_Tank_Value_Tank{0}_With_Filling_DryRun"
      on Click: InvertBit("DB702_Tank_Value_Tank{0}_With_Filling_DryRun")
   Button "Button_10" at 692,165 size 451x280; TextOff 'Text'
      Visibility <- "Control2"
   TextField "Text field_32" at 766,249 size 151x25; Text 'Tempering Unit'
      Visibility <- "Control2"
   TextField "Text field_33" at 766,296 size 163x25; Text 'Cool water valve'
      Visibility <- "Control2"
   TextField "Text field_34" at 766,343 size 141x25; Text 'Heater BackFL'
      Visibility <- "Control2"
   TextField "Text field_36" at 1002,296 size 68x25; Text 'Heater'
      Visibility <- "Control2"
   TextField "Text field_37" at 1002,343 size 129x25; Text 'Fischer valve'
      Visibility <- "Control2"
   TextField "Text field_38" at 719,194 size 232x30; Text 'Tempering Control :'
      Visibility <- "Control2"
   Button "Check_Tank_TC_TemperingUnit" at 711,246 size 45x30; TextOff 'Text'; PictureOff "download"; PictureList "Check_Uncheck"
      Visibility <- "Control2"
      on Click: InvertBit("DB702_Tank_Value_Tank{0}_With_Tempering_TempGeraet")
      ProcessValue <- "DB702_Tank_Value_Tank{0}_With_Tempering_TempGeraet"
   Button "Check_Tank_TC_CoolWaterValve" at 711,293 size 45x30; TextOff 'Text'; PictureOff "download"; PictureList "Check_Uncheck"
      Visibility <- "Control2"
      ProcessValue <- "DB702_Tank_Value_Tank{0}_With_Tempering_VKaltwasser"
      on Click: InvertBit("DB702_Tank_Value_Tank{0}_With_Tempering_VKaltwasser")
   Button "Check_Tank_TC_HeaterBackFL" at 711,340 size 45x30; TextOff 'Text'; PictureOff "download"; PictureList "Check_Uncheck"
      Visibility <- "Control2"
      on Click: InvertBit("DB702_Tank_Value_Tank{0}_With_Tempering_WTRL")
      ProcessValue <- "DB702_Tank_Value_Tank{0}_With_Tempering_WTRL"
   Button "Check_Tank_TC_Heater" at 948,293 size 45x30; TextOff 'Text'; PictureOff "download"; PictureList "Check_Uncheck"
      Visibility <- "Control2"
      ProcessValue <- "DB702_Tank_Value_Tank{0}_With_Tempering_Heizung"
      on Click: InvertBit("DB702_Tank_Value_Tank{0}_With_Tempering_Heizung")
   Button "Check_Tank_TC_FischerValve" at 948,340 size 45x30; TextOff 'Text'; PictureOff "download"; PictureList "Check_Uncheck"
      Visibility <- "Control2"
      ProcessValue <- "DB702_Tank_Value_Tank{0}_With_Tempering_WTmitFischer"
      on Click: InvertBit("DB702_Tank_Value_Tank{0}_With_Tempering_WTmitFischer")
   Button "b_Tank_Close_TemperingControl" at 1087,169 size 51x41; TextOff 'Text'; PictureOff "images (1)"
      Visibility <- "Control2"
      on Click: SetTag("Control2", 0)
   TextField "Text field_39" at 766,388 size 141x25; Text 'Heater Bypass'
      Visibility <- "Control2"
   Button "Check_Tank_HeaterBypass" at 711,385 size 45x30; TextOff 'Text'; PictureOff "download"; PictureList "Check_Uncheck"
      Visibility <- "Control2"
      ProcessValue <- "DB702_Tank_Value_Tank{0}_With_Tempering_WTBypass"
      on Click: InvertBit("DB702_Tank_Value_Tank{0}_With_Tempering_WTBypass")
   TextField "Text field_40" at 1002,389 size 128x25; Text 'Heater PreFl.'
      Visibility <- "Control2"
   Button "Check_Tank_TC_Heater_PreFL" at 948,386 size 45x30; TextOff 'Text'; PictureOff "download"; PictureList "Check_Uncheck"
      Visibility <- "Control2"
      ProcessValue <- "DB702_Tank_Value_Tank{0}_With_Tempering_WTVL"
      on Click: InvertBit("DB702_Tank_Value_Tank{0}_With_Tempering_WTVL")
   Button "BS POPUP" at 693,165 size 451x280; TextOff 'Text'
      Visibility <- "Control2"
   TextField "Text field_35" at 767,249 size 81x25; Text 'Existing'
      Visibility <- "Control2"
   TextField "Text field_41" at 767,296 size 94x25; Text 'pn. Pump'
      Visibility <- "Control2"
   TextField "Text field_42" at 767,343 size 102x25; Text 'pn. Stirrer'
      Visibility <- "Control2"
   TextField "Text field_43" at 1003,296 size 87x25; Text 'el. Pump'
      Visibility <- "Control2"
   TextField "Text field_44" at 1003,343 size 95x25; Text 'el. Stirrer'
      Visibility <- "Control2"
   TextField "Text field_45" at 712,194 size 171x30; Text 'Barrel station:'
      Visibility <- "Control2"
   Button "Check_Tank_BS_Existing" at 712,246 size 45x30; TextOff 'Text'; PictureOff "download"; PictureList "Check_Uncheck"
      Visibility <- "Control2"
      ProcessValue <- "DB702_Tank_Value_Tank{0}_With_BarelStation"
      on Click: InvertBit("DB702_Tank_Value_Tank{0}_With_BarelStation")
   Button "Check_Tank_BS_pnPump" at 712,293 size 45x30; TextOff 'Text'; PictureOff "download"; PictureList "Check_Uncheck"
      Visibility <- "Control2"
      ProcessValue <- "DB702_Tank_Value_Tank{0}_With_BarelStation_PnPump"
      on Click: InvertBit("DB702_Tank_Value_Tank{0}_With_BarelStation_PnPump")
   Button "Check_Tank_BS_pnStirrer" at 712,340 size 45x30; TextOff 'Text'; PictureOff "download"; PictureList "Check_Uncheck"
      Visibility <- "Control2"
      ProcessValue <- "DB702_Tank_Value_Tank{0}_With_BarelStation_PnRW"
      on Click: InvertBit("DB702_Tank_Value_Tank{0}_With_BarelStation_PnRW")
   Button "Check_Tank_BS_elPump" at 949,293 size 45x30; TextOff 'Text'; PictureOff "download"; PictureList "Check_Uncheck"
      Visibility <- "Control2"
      ProcessValue <- "DB702_Tank_Value_Tank{0}_With_BarelStation_ElPump"
      on Click: InvertBit("DB702_Tank_Value_Tank{0}_With_BarelStation_ElPump")
   Button "Check_Tank_BS_elStirrer" at 949,340 size 45x30; TextOff 'Text'; PictureOff "download"; PictureList "Check_Uncheck"
      Visibility <- "Control2"
      ProcessValue <- "DB702_Tank_Value_Tank{0}_With_BarelStation_ElRW"
      on Click: InvertBit("DB702_Tank_Value_Tank{0}_With_BarelStation_ElRW")
   Button "b_Tank_Close_BarrelStation" at 1088,169 size 51x41; TextOff 'Text'; PictureOff "images (1)"
      Visibility <- "Control2"
      on Click: SetTag("Control2", 0)
   TextField "Text field_46" at 767,389 size 116x25; Text 'Heat Jacket'
      Visibility <- "Control2"
   Button "Check_Tank_BS_HeatJacket" at 712,386 size 45x30; TextOff 'Text'; PictureOff "download"; PictureList "Check_Uncheck"
      Visibility <- "Control2"
      ProcessValue <- "DB702_Tank_Value_Tank{0}_With_BarelStation_Heating"
      on Click: InvertBit("DB702_Tank_Value_Tank{0}_With_BarelStation_Heating")
   TextField "Text field_47" at 1003,390 size 125x25; Text 'Heat Bottom'
      Visibility <- "Control2"
   Button "Check_Tank_BS_HeatBottom" at 949,387 size 45x30; TextOff 'Text'; PictureOff "download"; PictureList "Check_Uncheck"
      Visibility <- "Control2"
      ProcessValue <- "DB702_Tank_Value_Tank{0}_With_BarelStation_HeatingBottom"
      on Click: InvertBit("DB702_Tank_Value_Tank{0}_With_BarelStation_HeatingBottom")
   TextField "Text field_48" at 1004,251 size 108x25; Text 'Circulation'
      Visibility <- "Control2"
   Button "Check_Tank_BS_Circulation" at 950,248 size 45x30; TextOff 'Text'; PictureOff "download"; PictureList "Check_Uncheck"
      Visibility <- "Control2"
      ProcessValue <- "DB702_Tank_Value_Tank{0}_With_BarelStation_Zirkulation"
      on Click: InvertBit("DB702_Tank_Value_Tank{0}_With_BarelStation_Zirkulation")
   Button "Stirrer POPUP" at 693,164 size 451x280; TextOff 'Text'
      Visibility <- "Control2"
   TextField "Text field_49" at 767,248 size 81x25; Text 'Existing'
      Visibility <- "Control2"
   TextField "Text field_50" at 767,295 size 98x25; Text 'Converter'
      Visibility <- "Control2"
   TextField "Text field_51" at 767,342 size 94x25; Text 'Set Value'
      Visibility <- "Control2"
   TextField "Text field_53" at 1003,342 size 112x25; Text '6 Set Value'
      Visibility <- "Control2"
   TextField "Text field_54" at 712,193 size 88x30; Text 'Stirrer:'
      Visibility <- "Control2"
   Button "Check_Tank_Stirrer_Existing" at 712,245 size 45x30; TextOff 'Text'; PictureOff "download"; PictureList "Check_Uncheck"
      Visibility <- "Control2"
      on Click: InvertBit("DB702_Tank_Value_Tank{0}_With_Agitator")
      ProcessValue <- "DB702_Tank_Value_Tank{0}_With_Agitator"
   Button "Check_Tank_Stirrer_Converter" at 712,292 size 45x30; TextOff 'Text'; PictureOff "download"; PictureList "Check_Uncheck"
      Visibility <- "Control2"
      on Click: InvertBit("DB702_Tank_Value_Tank{0}_With_Agitator_Converter")
      ProcessValue <- "DB702_Tank_Value_Tank{0}_With_Agitator_Converter"
   Button "Check_Tank_Stirrer_SetValue" at 712,339 size 45x30; TextOff 'Text'; PictureOff "download"; PictureList "Check_Uncheck"
      Visibility <- "Control2"
      ProcessValue <- "DB702_Tank_Value_Tank{0}_With_Agitator_SetValue"
      on Click: InvertBit("DB702_Tank_Value_Tank{0}_With_Agitator_SetValue")
   Button "Check_Tank_Stirrer_6SetValue" at 949,339 size 45x30; TextOff 'Text'; PictureOff "download"; PictureList "Check_Uncheck"
      Visibility <- "Control2"
      ProcessValue <- "DB702_Tank_Value_Tank{0}_With_Agitator_6SetValue"
      on Click: InvertBit("DB702_Tank_Value_Tank{0}_With_Agitator_6SetValue")
   Button "b_Tank_Close_Strirrer" at 1088,168 size 51x41; TextOff 'Text'; PictureOff "images (1)"
      on Press: SetTag("Control2", 0)
      Visibility <- "Control2"
   Button "ForceStirring POPUP" at 693,163 size 451x280; TextOff 'Text'
      Visibility <- "Control2"
   TextField "Text field_52" at 767,247 size 79x25; Text 'Heating'
      Visibility <- "Control2"
   TextField "Text field_55" at 767,294 size 77x25; Text 'Cooling'
      Visibility <- "Control2"
   TextField "Text field_56" at 767,341 size 64x25; Text 'Filling'
      Visibility <- "Control2"
   TextField "Text field_57" at 1003,294 size 81x25; Text 'Interval'
      Visibility <- "Control2"
   TextField "Text field_58" at 1003,341 size 81x25; Text 'Interval'
      Visibility <- "Control2"
   TextField "Text field_59" at 712,192 size 169x30; Text 'Force Stirring:'
      Visibility <- "Control2"
   Button "Check_Tank_FS_Heating" at 712,244 size 45x30; TextOff 'Text'; PictureOff "download"; PictureList "Check_Uncheck"
      Visibility <- "Control2"
      on Click: InvertBit("DB702_Tank_Value_Tank{0}_Agitator_Config_bit_Heating_ON")
      ProcessValue <- "DB702_Tank_Value_Tank{0}_Agitator_Config_bit_Heating_ON"
   Button "Check_Tank_FS_Cooling" at 712,291 size 45x30; TextOff 'Text'; PictureOff "download"; PictureList "Check_Uncheck"
      Visibility <- "Control2"
      on Click: InvertBit("DB702_Tank_Value_Tank{0}_Agitator_Config_bit_Cooling_ON")
      ProcessValue <- "DB702_Tank_Value_Tank{0}_Agitator_Config_bit_Cooling_ON"
   Button "Check_Tank_FS_Filling" at 712,338 size 45x30; TextOff 'Text'; PictureOff "download"; PictureList "Check_Uncheck"
      Visibility <- "Control2"
      on Click: InvertBit("DB702_Tank_Value_Tank{0}_Agitator_Config_bit_Filling_ON")
      ProcessValue <- "DB702_Tank_Value_Tank{0}_Agitator_Config_bit_Filling_ON"
   Button "Check_Tank_FS_Interval2" at 949,291 size 45x30; TextOff 'Text'; PictureOff "download"; PictureList "Check_Uncheck"
      Visibility <- "Control2"
      on Click: InvertBit("DB702_Tank_Value_Tank{0}_Agitator_Config_bit_Cooling_Int")
      ProcessValue <- "DB702_Tank_Value_Tank{0}_Agitator_Config_bit_Cooling_Int"
   Button "Check_Tank_FS_Interval3" at 949,338 size 45x30; TextOff 'Text'; PictureOff "download"; PictureList "Check_Uncheck"
      Visibility <- "Control2"
      on Click: InvertBit("DB702_Tank_Value_Tank{0}_Agitator_Config_bit_Filling_Int")
      ProcessValue <- "DB702_Tank_Value_Tank{0}_Agitator_Config_bit_Filling_Int"
   Button "b_Tank_Close_ForceStrirring" at 1088,167 size 51x41; TextOff 'Text'; PictureOff "images (1)"
      on Press: SetTag("Control2", 0)
      Visibility <- "Control2"
   TextField "Text field_60" at 767,386 size 108x25; Text 'Taking Out'
      Visibility <- "Control2"
   Button "Check_Tank_FS_TakingOut" at 712,383 size 45x30; TextOff 'Text'; PictureOff "download"; PictureList "Check_Uncheck"
      Visibility <- "Control2"
      on Click: InvertBit("DB702_Tank_Value_Tank{0}_Agitator_Config_bit_Charging_ON")
      ProcessValue <- "DB702_Tank_Value_Tank{0}_Agitator_Config_bit_Charging_ON"
   TextField "Text field_61" at 1003,387 size 81x25; Text 'Interval'
      Visibility <- "Control2"
   Button "Check_Tank_FS_Interval4" at 949,384 size 45x30; TextOff 'Text'; PictureOff "download"; PictureList "Check_Uncheck"
      Visibility <- "Control2"
      on Click: InvertBit("DB702_Tank_Value_Tank{0}_Agitator_Config_bit_Charging_Int")
      ProcessValue <- "DB702_Tank_Value_Tank{0}_Agitator_Config_bit_Charging_Int"
   TextField "Text field_62" at 1004,249 size 81x25; Text 'Interval'
      Visibility <- "Control2"
   Button "Check_Tank_FS_Interval1" at 950,246 size 45x30; TextOff 'Text'; PictureOff "download"; PictureList "Check_Uncheck"
      Visibility <- "Control2"
      on Click: InvertBit("DB702_Tank_Value_Tank{0}_Agitator_config_bit_Heating_Int")
      ProcessValue <- "DB702_Tank_Value_Tank{0}_Agitator_config_bit_Heating_Int"
   Button "Button_3" at 116,166 size 535x569; TextOff 'Text'; PictureOff "tank"
      Visibility <- "DB702_Tank_Value_Tank{0}_Existing"
      on Press: InvertBit("DB702_Tank_Value_Tank{0}_Existing")
   Rectangle "Rectangle_4" at 147,608 size 456x40
      Visibility <- "DB702_Tank_Value_Tank{0}_With_Agitator"